REGION Network 9: No encoder pulse
   RUNG wire#powerrail
      Contact( #IN_xFaultsEnabled )
      Contact( #IN_xCycleONDel )
      Contact( #ST_xEncDownPosition )
      { S7_Templates := "SrcType := DInt" } EQ_Contact(in1 := #INPUTS.dEncCounter_count, in2 := #AUX_dLastCounterValueFast_cmm)
      Move(in := #INPUTS.dEncCounter_count, out1 => #AUX_dLastCounterValueFast_cmm)
      Coil( #tALM.tS.xNoEncPulses )
   END_RUNG
   // the same network as SCL:
   #_w1 := #IN_xFaultsEnabled AND #IN_xCycleONDel AND #ST_xEncDownPosition AND (#INPUTS.dEncCounter_count = #AUX_dLastCounterValueFast_cmm);
   IF #_w1 THEN #AUX_dLastCounterValueFast_cmm := #INPUTS.dEncCounter_count; END_IF;
   #tALM.tS.xNoEncPulses := #_w1;
END_REGION

REGION Network 10: Speed values outside limits
   RUNG wire#powerrail
      Contact( #IN_xFaultsEnabled )
      Contact( #IN_xCycleONDel )
      Contact( #ST_xEncDownPosition )
      wire#w1
      { S7_Templates := "SrcType := DInt" } LT_Contact(in1 := #tHMR.dActualEncoderSpeed_mm_min, in2 := "DMINLEHRSPEED_MM_MIN")
      wire#w2
      Coil( #tALM.tS.xSpeedOutLimits )
   END_RUNG
   RUNG wire#w1
      { S7_Templates := "SrcType := DInt" } GT_Contact(in1 := #tHMR.dActualEncoderSpeed_mm_min, in2 := "DMAXLEHRSPEED_MM_MIN")
   END_RUNG wire#w2
   // the same network as SCL:
   #tALM.tS.xSpeedOutLimits := #IN_xFaultsEnabled AND #IN_xCycleONDel AND #ST_xEncDownPosition AND ((#tHMR.dActualEncoderSpeed_mm_min < "DMINLEHRSPEED_MM_MIN") OR (#tHMR.dActualEncoderSpeed_mm_min > "DMAXLEHRSPEED_MM_MIN"));
END_REGION

REGION Network 11: Fm152. Sending data error
   RUNG wire#powerrail
      Contact( #tPhases.xEndPrepareTelegram )
      Contact( #FB_TSend.ERROR )
      S_Coil( #tALM.tF.xFm152SendError )
   END_RUNG
   // the same network as SCL:
   IF #tPhases.xEndPrepareTelegram AND #FB_TSend.ERROR THEN #tALM.tF.xFm152SendError := TRUE; END_IF;
END_REGION

REGION Network 12: FM152.Send data timeout
   #tmON_TimeoutSendData(IN := #tPhases.xPrepareTelegram, PT := #CONST_DTIMEOUTSENDDATA_MS);   // TON
   IF #tmON_TimeoutSendData.Q THEN #tALM.tF.xFm152SendTimeout := TRUE; END_IF;
END_REGION

REGION Network 13: Receive timeout
   #tmON_TimeoutRecvData(IN := #tPhases.xWaitingFm152Reply, PT := #CONST_DTIMEOUTRECVDATA_MS);   // TON
   IF #tmON_TimeoutRecvData.Q THEN
       #tALM.tF.xFm152RecvTimeout := TRUE;
       #AUX_dActualElBuffer := 0;
   END_IF;
END_REGION

REGION Network 14 (SCL): Calculate general statuses
   GATHER(IN:=#tALM.tS,
          OUT=>#TMP_dwValue);

   IF #TMP_dwValue <> 0 THEN
       #ST_xStoppingFaults := TRUE;
   ELSE
       #ST_xStoppingFaults := FALSE;
   END_IF;

   GATHER(IN:=#tALM.tF,
          OUT=>#TMP_dwValue);

   IF #TMP_dwValue <> 0 THEN
       #ST_xFaults := TRUE;
   ELSE
       #ST_xFaults := FALSE;
   END_IF;

   GATHER(IN:=#tALM.tW,
          OUT=>#TMP_dwValue);

   IF #TMP_dwValue <> 0 THEN
       #ST_xWarnings := TRUE;
   ELSE
       #ST_xWarnings := FALSE;
   END_IF;
END_REGION

REGION Network 15: ####_HMI_LOGICS_####
END_REGION

REGION Network 16 (SCL): Manage HMI request
   (*REGION Enable disable glass sensor

       IF #tHMW.xEnableGlassSensor THEN
           #tHMR.xGlassSensorEnabled := TRUE;
           #tHMW.xEnableGlassSensor := FALSE;
       END_IF;

       IF #tHMW.xDisableGlassSensor THEN
           #tHMR.xGlassSensorEnabled := FALSE;
           #tHMW.xDisableGlassSensor := FALSE;
       END_IF;

   END_REGION *)

   REGION Length calibration

       IF #tHMW.xCalibRequest THEN

           #TMP_rF1Unit := DINT_TO_REAL(#tHMW.dCalibRealLength_cmm) / (DINT_TO_REAL(#tHMW.dCalibTheoLength_cmm) / DINT_TO_REAL(#tHMR.dCalibrationF1Unit_unit));
           #tHMR.dCalibrationF1Unit_unit := REAL_TO_DINT(#TMP_rF1Unit);

           #tHMW.dCalibRealLength_cmm := #tHMW.dCalibTheoLength_cmm;        

           #tHMW.xCalibRequest := FALSE;

       END_IF;

   END_REGION

   REGION Update F1

       IF #tHMW.xCalibUpdateF1 THEN

           #tHMR.dCalibrationF1Unit_unit := #tHMW.dCalibWriteF1_unit;
           #tHMW.xCalibUpdateF1 := FALSE;
           #ST_xRefreshFM152 := TRUE;

       END_IF;

   END_REGION

   REGION Update F2

       IF #tHMW.xCalibUpdateF2 THEN

           #tHMR.dCalibrationF2Unit_unit := #tHMW.dCalibWriteF2_unit;
           #tHMW.xCalibUpdateF2 := FALSE;
           #ST_xRefreshFM152 := TRUE;

       END_IF;

   END_REGION
END_REGION

REGION Network 17: Manual command enabled
   RUNG wire#powerrail
      Contact( #tHMW.xEnDisManCom )
      Contact( #ST_xCondOkMan )
      wire#w1
      Coil( #tHMR.xManComEn )
   END_RUNG
   RUNG wire#powerrail
      Contact( #tHMR.xManComEn )
      Contact( #tHMW.xEnDisManCom )
   END_RUNG wire#w1
   // the same network as SCL:
   #tHMR.xManComEn := (#tHMW.xEnDisManCom AND #ST_xCondOkMan) OR (#tHMR.xManComEn AND #tHMW.xEnDisManCom);
END_REGION

REGION Network 18: ####_STATUSES_####
END_REGION

REGION Network 19: Output enable
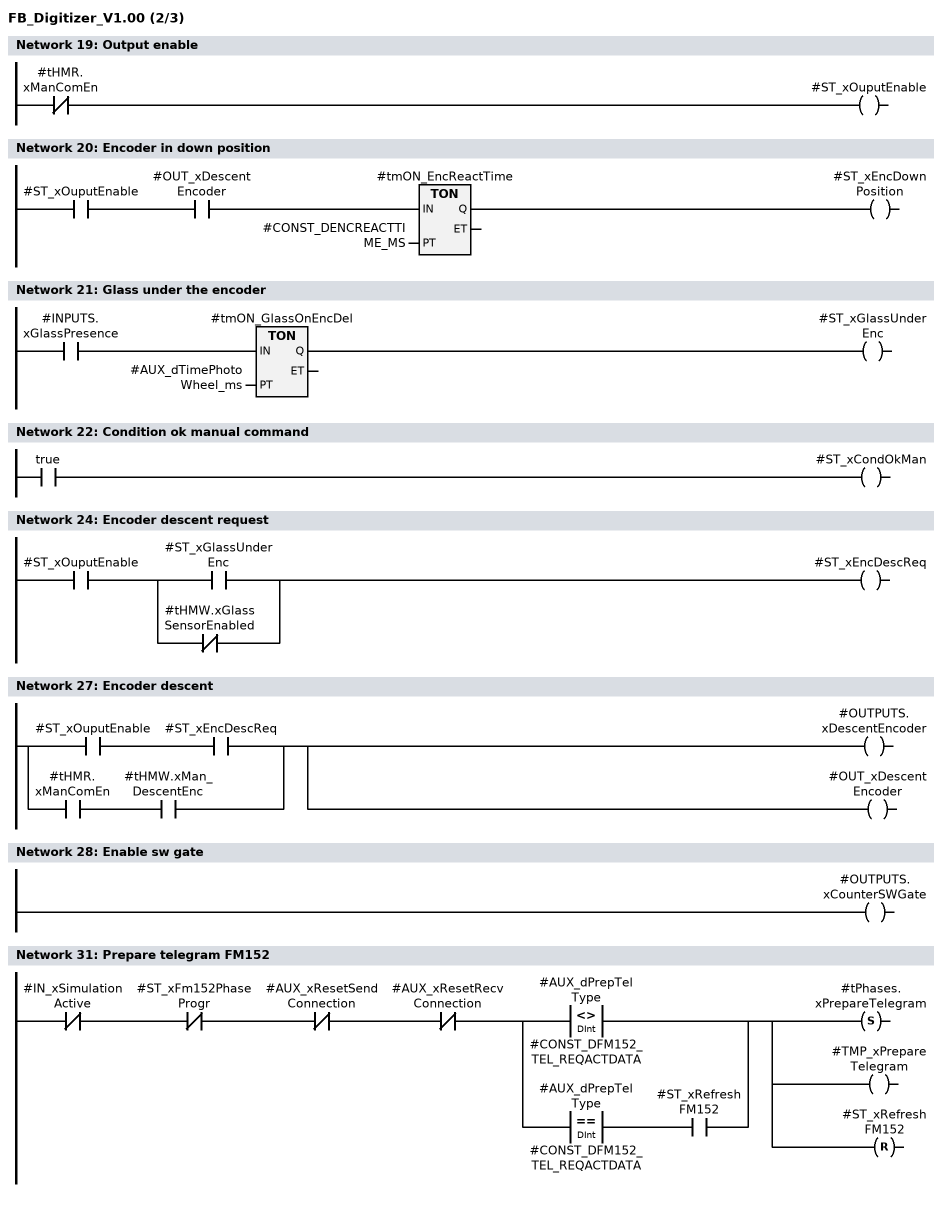
   RUNG wire#powerrail
      I_Contact( #tHMR.xManComEn )
      Coil( #ST_xOuputEnable )
   END_RUNG
   // the same network as SCL:
   #ST_xOuputEnable := NOT #tHMR.xManComEn;
END_REGION

REGION Network 20: Encoder in down position
   #tmON_EncReactTime(IN := #ST_xOuputEnable AND #OUT_xDescentEncoder, PT := #CONST_DENCREACTTIME_MS);   // TON
   #ST_xEncDownPosition := #tmON_EncReactTime.Q;
END_REGION

REGION Network 21: Glass under the encoder
   #tmON_GlassOnEncDel(IN := #INPUTS.xGlassPresence, PT := #AUX_dTimePhotoWheel_ms);   // TON
   #ST_xGlassUnderEnc := #tmON_GlassOnEncDel.Q;
END_REGION

REGION Network 22: Condition ok manual command
   RUNG wire#powerrail
      Contact( true )
      Coil( #ST_xCondOkMan )
   END_RUNG
   // the same network as SCL:
   #ST_xCondOkMan := true;
END_REGION

REGION Network 23: ####_PHASES_&_LOGICS_####
END_REGION

REGION Network 24: Encoder descent request
   RUNG wire#powerrail
      Contact( #ST_xOuputEnable )
      wire#w1
      Contact( #ST_xGlassUnderEnc )
      wire#w2
      Coil( #ST_xEncDescReq )
   END_RUNG
   RUNG wire#w1
      I_Contact( #tHMW.xGlassSensorEnabled )
   END_RUNG wire#w2
   // the same network as SCL:
   #ST_xEncDescReq := #ST_xOuputEnable AND (#ST_xGlassUnderEnc OR NOT #tHMW.xGlassSensorEnabled);
END_REGION

REGION Network 25 (SCL): ####_HMI_STATUSES_####
   #AUX_lrTimingCounter_s += #AUX_lrElapsedTime_s;

   IF #AUX_lrTimingCounter_s >= #CONST_DREFRESHSPEED_S THEN

       #TMP_dElapsedPulses_cmm := #INPUTS.dEncCounter_count - #AUX_dLastCounterValue_cmm;

       #tHMR.dActualEncoderSpeed_mm_min := REAL_TO_DINT(((DINT_TO_REAL(#TMP_dElapsedPulses_cmm) / 100.0) / (LREAL_TO_REAL(#AUX_lrTimingCounter_s))) * 60.0);

       #AUX_dLastCounterValue_cmm := #INPUTS.dEncCounter_count;
       #AUX_lrTimingCounter_s := 0;

   END_IF;

   IF #OUTPUTS.xDescentEncoder AND #tHMW.xMan_DescentEnc THEN
       #tHMR.xMan_DescEncFdbk := TRUE;
   ELSE
       #tHMR.xMan_DescEncFdbk := FALSE;

   END_IF;

   IF #ST_xStoppingFaults THEN
       #tHMR.dEncoderStatus := 7;
   ELSIF #ST_xEncDownPosition THEN
       #tHMR.dEncoderStatus := 3;
   ELSE
       #tHMR.dEncoderStatus := 1;
   END_IF;
END_REGION

REGION Network 26: ####_OUTPUTS_####
END_REGION

REGION Network 27: Encoder descent
   RUNG wire#powerrail
      Contact( #ST_xOuputEnable )
      Contact( #ST_xEncDescReq )
      wire#w1
      Coil( #OUTPUTS.xDescentEncoder )
   END_RUNG
   RUNG wire#powerrail
      Contact( #tHMR.xManComEn )
      Contact( #tHMW.xMan_DescentEnc )
   END_RUNG wire#w1
   RUNG wire#w1
      Coil( #OUT_xDescentEncoder )
   END_RUNG
   // the same network as SCL:
   #OUTPUTS.xDescentEncoder := (#ST_xOuputEnable AND #ST_xEncDescReq) OR (#tHMR.xManComEn AND #tHMW.xMan_DescentEnc);
   #OUT_xDescentEncoder := #OUTPUTS.xDescentEncoder;
END_REGION

REGION Network 28: Enable sw gate
   RUNG wire#powerrail
      Coil( #OUTPUTS.xCounterSWGate )
   END_RUNG
   // the same network as SCL:
   #OUTPUTS.xCounterSWGate := TRUE;
END_REGION

REGION Network 29: ####_ETHERNET_TO_FM152_####
END_REGION

REGION Network 30 (SCL): Initialize connection data
   IF #IN_xGeneralReset THEN

       #AUX_tConnData.InterfaceId := #IN_tInterfaceID;
       #AUX_tConnData.ID := #IN_tID;
       #AUX_tConnData.ConnectionType := #CONST_BCONNTYPE;
       #AUX_tConnData.ActiveEstablished := TRUE;
       #AUX_tConnData.RemoteAddress := #IN_tRemoteAddress;
       #AUX_tConnData.RemotePort := #IN_uiRemotePort;
       #AUX_tConnData.LocalPort := 0;

       //Reset della fasi
       #TMP_dwValue := 0;
       SCATTER(IN:=#TMP_dwValue,
               OUT=>#tPhases);



   END_IF;

   #AUX_xResetRecvConnection := #IN_xGeneralReset;
   #AUX_xResetSendConnection := #IN_xGeneralReset;
END_REGION

REGION Network 31: Prepare telegram FM152
   RUNG wire#powerrail
      I_Contact( #IN_xSimulationActive )
      I_Contact( #ST_xFm152PhaseProgr )
      I_Contact( #AUX_xResetSendConnection )
      I_Contact( #AUX_xResetRecvConnection )
      wire#w1
      { S7_Templates := "SrcType := DInt" } NE_Contact(in1 := #AUX_dPrepTelType, in2 := #CONST_DFM152_TEL_REQACTDATA)
      wire#w2
      S_Coil( #tPhases.xPrepareTelegram )
   END_RUNG
   RUNG wire#w1
      { S7_Templates := "SrcType := DInt" } EQ_Contact(in1 := #AUX_dPrepTelType, in2 := #CONST_DFM152_TEL_REQACTDATA)
      Contact( #ST_xRefreshFM152 )
   END_RUNG wire#w2
   RUNG wire#w2
      Coil( #TMP_xPrepareTelegram )
   END_RUNG
   RUNG wire#w2
      R_Coil( #ST_xRefreshFM152 )
   END_RUNG
   // the same network as SCL:
   #_w1 := NOT #IN_xSimulationActive AND NOT #ST_xFm152PhaseProgr AND NOT #AUX_xResetSendConnection AND NOT #AUX_xResetRecvConnection AND ((#AUX_dPrepTelType <> #CONST_DFM152_TEL_REQACTDATA) OR ((#AUX_dPrepTelType = #CONST_DFM152_TEL_REQACTDATA) AND #ST_xRefreshFM152));
   IF #_w1 THEN #tPhases.xPrepareTelegram := TRUE; END_IF;
   #TMP_xPrepareTelegram := #_w1;
   IF #_w1 THEN #ST_xRefreshFM152 := FALSE; END_IF;
END_REGION

REGION Network 32 (SCL): Prepare telegram
   IF #TMP_xPrepareTelegram THEN

       #AUX_dPrepTelType += 1;

       IF #AUX_dPrepTelType > #CONST_DFM152_TEL_REQACTDATA THEN
           #AUX_dPrepTelType := #CONST_DFM152_TEL_READST;
       END_IF;

       CASE #AUX_dPrepTelType OF

           #CONST_DFM152_TEL_READST:

               #AUX_tFM152SndReadSt.bEOT := #CONST_BFM152_EOT;
               #AUX_tFM152SndReadSt.bAD1 := #CONST_BFM152_AD1;    
               #AUX_tFM152SndReadSt.bAD2 := #CONST_BFM152_AD2;
               #AUX_tFM152SndReadSt.bC1 := '8';
               #AUX_tFM152SndReadSt.bC2 := '5';
               #AUX_tFM152SndReadSt.bENQ := #CONST_BFM152_ENQ;

               #TMP_dBufferPos := 0;
               #TMP_iRetVal := Serialize(SRC_VARIABLE:=#AUX_tFM152SndReadSt, DEST_ARRAY=>#AUX_rgbTempSendBuffer, POS:=#TMP_dBufferPos);
               #AUX_dNumByteToSend := #CONST_DFM152_TEL_READST_NUMBYTE;

           #CONST_DFM152_TEL_READF1:

               #AUX_tFM152SndReadF1.bEOT := #CONST_BFM152_EOT;
               #AUX_tFM152SndReadF1.bAD1 := #CONST_BFM152_AD1;    
               #AUX_tFM152SndReadF1.bAD2 := #CONST_BFM152_AD2;
               #AUX_tFM152SndReadF1.bC1 := '0';
               #AUX_tFM152SndReadF1.bC2 := '0';
               #AUX_tFM152SndReadF1.bENQ := #CONST_BFM152_ENQ;

               #TMP_dBufferPos := 0;
               #TMP_iRetVal := Serialize(SRC_VARIABLE:=#AUX_tFM152SndReadF1, DEST_ARRAY=>#AUX_rgbTempSendBuffer, POS:=#TMP_dBufferPos);
               #AUX_dNumByteToSend := #CONST_DFM152_TEL_READF1_NUMBYTE;

           #CONST_DFM152_TEL_READF2:

               #AUX_tFM152SndReadF2.bEOT := #CONST_BFM152_EOT;
               #AUX_tFM152SndReadF2.bAD1 := #CONST_BFM152_AD1;    
               #AUX_tFM152SndReadF2.bAD2 := #CONST_BFM152_AD2;
               #AUX_tFM152SndReadF2.bC1 := '0';
               #AUX_tFM152SndReadF2.bC2 := '1';
               #AUX_tFM152SndReadF2.bENQ := #CONST_BFM152_ENQ;

               #TMP_dBufferPos := 0;
               #TMP_iRetVal := Serialize(SRC_VARIABLE:=#AUX_tFM152SndReadF2, DEST_ARRAY=>#AUX_rgbTempSendBuffer, POS:=#TMP_dBufferPos);
               #AUX_dNumByteToSend := #CONST_DFM152_TEL_READF2_NUMBYTE;

           #CONST_DFM152_TEL_WRITEF1:

               #TMP_strValue := DINT_TO_STRING(#tHMR.dCalibrationF1Unit_unit);

               #AUX_tFM152SndWriteF1.bEOT := #CONST_BFM152_EOT;
               #AUX_tFM152SndWriteF1.bAD1 := #CONST_BFM152_AD1;
               #AUX_tFM152SndWriteF1.bAD2 := #CONST_BFM152_AD2;
               #AUX_tFM152SndWriteF1.bSTX := #CONST_BFM152_STX;
               #AUX_tFM152SndWriteF1.bC1 := '0';
               #AUX_tFM152SndWriteF1.bC2 := '0';
               #AUX_tFM152SndWriteF1.bVal1 := #TMP_strValue[2];
               #AUX_tFM152SndWriteF1.bVal2 := #TMP_strValue[3];
               #AUX_tFM152SndWriteF1.bVal3 := #TMP_strValue[4];
               #AUX_tFM152SndWriteF1.bVal4 := #TMP_strValue[5];
               #AUX_tFM152SndWriteF1.bVal5 := #TMP_strValue[6];
               #AUX_tFM152SndWriteF1.bETX := #CONST_BFM152_ETX;
               #AUX_tFM152SndWriteF1.bBCC := #AUX_tFM152SndWriteF1.bC1; 
               #AUX_tFM152SndWriteF1.bBCC := #AUX_tFM152SndWriteF1.bBCC XOR #AUX_tFM152SndWriteF1.bC2;
               #AUX_tFM152SndWriteF1.bBCC := #AUX_tFM152SndWriteF1.bBCC XOR #AUX_tFM152SndWriteF1.bVal1;
               #AUX_tFM152SndWriteF1.bBCC := #AUX_tFM152SndWriteF1.bBCC XOR #AUX_tFM152SndWriteF1.bVal2;
               #AUX_tFM152SndWriteF1.bBCC := #AUX_tFM152SndWriteF1.bBCC XOR #AUX_tFM152SndWriteF1.bVal3;
               #AUX_tFM152SndWriteF1.bBCC := #AUX_tFM152SndWriteF1.bBCC XOR #AUX_tFM152SndWriteF1.bVal4;
               #AUX_tFM152SndWriteF1.bBCC := #AUX_tFM152SndWriteF1.bBCC XOR #AUX_tFM152SndWriteF1.bVal5;
               #AUX_tFM152SndWriteF1.bBCC := #AUX_tFM152SndWriteF1.bBCC XOR #AUX_tFM152SndWriteF1.bETX; 

               #TMP_dBufferPos := 0;
               #TMP_iRetVal := Serialize(SRC_VARIABLE:=#AUX_tFM152SndWriteF1, DEST_ARRAY=>#AUX_rgbTempSendBuffer, POS:=#TMP_dBufferPos);
               #AUX_dNumByteToSend := #CONST_DFM152_TEL_WRITEF1_NUMBYTE;

           #CONST_DFM152_TEL_WRITEF2:

               #TMP_strValue := DINT_TO_STRING(#tHMR.dCalibrationF2Unit_unit);

               #AUX_tFM152SndWriteF2.bEOT := #CONST_BFM152_EOT;
               #AUX_tFM152SndWriteF2.bAD1 := #CONST_BFM152_AD1;
               #AUX_tFM152SndWriteF2.bAD2 := #CONST_BFM152_AD2;
               #AUX_tFM152SndWriteF2.bSTX := #CONST_BFM152_STX;
               #AUX_tFM152SndWriteF2.bC1 := '0';
               #AUX_tFM152SndWriteF2.bC2 := '1';
               #AUX_tFM152SndWriteF2.bVal1 := #TMP_strValue[2];
               #AUX_tFM152SndWriteF2.bVal2 := #TMP_strValue[3];
               #AUX_tFM152SndWriteF2.bVal3 := #TMP_strValue[4];
               #AUX_tFM152SndWriteF2.bVal4 := #TMP_strValue[5];
               #AUX_tFM152SndWriteF2.bVal5 := #TMP_strValue[6];
               #AUX_tFM152SndWriteF2.bETX := #CONST_BFM152_ETX;
               #AUX_tFM152SndWriteF2.bBCC := #AUX_tFM152SndWriteF2.bC1; 
               #AUX_tFM152SndWriteF2.bBCC := #AUX_tFM152SndWriteF2.bBCC XOR #AUX_tFM152SndWriteF2.bC2;
               #AUX_tFM152SndWriteF2.bBCC := #AUX_tFM152SndWriteF2.bBCC XOR #AUX_tFM152SndWriteF2.bVal1;
               #AUX_tFM152SndWriteF2.bBCC := #AUX_tFM152SndWriteF2.bBCC XOR #AUX_tFM152SndWriteF2.bVal2;
               #AUX_tFM152SndWriteF2.bBCC := #AUX_tFM152SndWriteF2.bBCC XOR #AUX_tFM152SndWriteF2.bVal3;
               #AUX_tFM152SndWriteF2.bBCC := #AUX_tFM152SndWriteF2.bBCC XOR #AUX_tFM152SndWriteF2.bVal4;
               #AUX_tFM152SndWriteF2.bBCC := #AUX_tFM152SndWriteF2.bBCC XOR #AUX_tFM152SndWriteF2.bVal5;
               #AUX_tFM152SndWriteF2.bBCC := #AUX_tFM152SndWriteF2.bBCC XOR #AUX_tFM152SndWriteF2.bETX; 

               #TMP_dBufferPos := 0;
               #TMP_iRetVal := Serialize(SRC_VARIABLE:=#AUX_tFM152SndWriteF2, DEST_ARRAY=>#AUX_rgbTempSendBuffer, POS:=#TMP_dBufferPos);
               #AUX_dNumByteToSend := #CONST_DFM152_TEL_WRITEF2_NUMBYTE;

           #CONST_DFM152_TEL_WRITEJOG:

               #TMP_strValue := DINT_TO_STRING(REAL_TO_DINT((DINT_TO_REAL(#tHMW.dRequestJogSpeed_mm_min) * 100.0) / 60.0));
               #AUX_tFM152SndWriteJog.bEOT := #CONST_BFM152_EOT;
               #AUX_tFM152SndWriteJog.bAD1 := #CONST_BFM152_AD1;
               #AUX_tFM152SndWriteJog.bAD2 :=  #CONST_BFM152_AD2;
               #AUX_tFM152SndWriteJog.bSTX := #CONST_BFM152_STX;
               #AUX_tFM152SndWriteJog.bC1 := '0'; 
               #AUX_tFM152SndWriteJog.bC2 := '5'; 
               #AUX_tFM152SndWriteJog.bVal1 := #TMP_strValue[2];
               #AUX_tFM152SndWriteJog.bVal2 := #TMP_strValue[3];
               #AUX_tFM152SndWriteJog.bVal3 := #TMP_strValue[4];
               #AUX_tFM152SndWriteJog.bVal4 := #TMP_strValue[5];
               #AUX_tFM152SndWriteJog.bVal5 := #TMP_strValue[6];
               #AUX_tFM152SndWriteJog.bETX := #CONST_BFM152_ETX;
               #AUX_tFM152SndWriteJog.bBCC := #AUX_tFM152SndWriteJog.bC1; 
               #AUX_tFM152SndWriteJog.bBCC := #AUX_tFM152SndWriteJog.bBCC XOR #AUX_tFM152SndWriteJog.bC2;
               #AUX_tFM152SndWriteJog.bBCC := #AUX_tFM152SndWriteJog.bBCC XOR #AUX_tFM152SndWriteJog.bVal1;
               #AUX_tFM152SndWriteJog.bBCC := #AUX_tFM152SndWriteJog.bBCC XOR #AUX_tFM152SndWriteJog.bVal2;
               #AUX_tFM152SndWriteJog.bBCC := #AUX_tFM152SndWriteJog.bBCC XOR #AUX_tFM152SndWriteJog.bVal3;
               #AUX_tFM152SndWriteJog.bBCC := #AUX_tFM152SndWriteJog.bBCC XOR #AUX_tFM152SndWriteJog.bVal4;
               #AUX_tFM152SndWriteJog.bBCC := #AUX_tFM152SndWriteJog.bBCC XOR #AUX_tFM152SndWriteJog.bVal5;
               #AUX_tFM152SndWriteJog.bBCC := #AUX_tFM152SndWriteJog.bBCC XOR #AUX_tFM152SndWriteJog.bETX;

               #TMP_dBufferPos := 0;
               #TMP_iRetVal := Serialize(SRC_VARIABLE:=#AUX_tFM152SndWriteJog, DEST_ARRAY=>#AUX_rgbTempSendBuffer, POS:=#TMP_dBufferPos);
               #AUX_dNumByteToSend := #CONST_DFM152_TEL_WRITEJOG_NUMBYTE;


           #CONST_DFM152_TEL_WRITERAMPREF:

               #AUX_tFM152SndWriteRampRef.bEOT := #CONST_BFM152_EOT;
               #AUX_tFM152SndWriteRampRef.bAD1 := #CONST_BFM152_AD1;
               #AUX_tFM152SndWriteRampRef.bAD2 := #CONST_BFM152_AD2;
               #AUX_tFM152SndWriteRampRef.bSTX := #CONST_BFM152_STX;
               #AUX_tFM152SndWriteRampRef.bC1 := '0';
               #AUX_tFM152SndWriteRampRef.bC2 := '4';
               #AUX_tFM152SndWriteRampRef.bC3 := '0';
               #AUX_tFM152SndWriteRampRef.bC4 := '0';
               #AUX_tFM152SndWriteRampRef.bETX := #CONST_BFM152_ETX;
               #AUX_tFM152SndWriteRampRef.bBCC := #AUX_tFM152SndWriteRampRef.bC1;
               #AUX_tFM152SndWriteRampRef.bBCC :=  #AUX_tFM152SndWriteRampRef.bBCC XOR #AUX_tFM152SndWriteRampRef.bC2;
               #AUX_tFM152SndWriteRampRef.bBCC :=  #AUX_tFM152SndWriteRampRef.bBCC XOR #AUX_tFM152SndWriteRampRef.bC3;
               #AUX_tFM152SndWriteRampRef.bBCC :=  #AUX_tFM152SndWriteRampRef.bBCC XOR #AUX_tFM152SndWriteRampRef.bC4;
               #AUX_tFM152SndWriteRampRef.bBCC :=  #AUX_tFM152SndWriteRampRef.bBCC XOR #AUX_tFM152SndWriteRampRef.bETX;

               #TMP_dBufferPos := 0;
               #TMP_iRetVal := Serialize(SRC_VARIABLE:=#AUX_tFM152SndWriteRampRef, DEST_ARRAY=>#AUX_rgbTempSendBuffer, POS:=#TMP_dBufferPos);
               #AUX_dNumByteToSend := #CONST_DFM152_TEL_WRITERAMPREF_NUMBYTE;


           #CONST_DFM152_TEL_WRITERAMPJOG:

               #AUX_tFM152SndWriteRampJog.bEOT := #CONST_BFM152_EOT;
               #AUX_tFM152SndWriteRampJog.bAD1 := #CONST_BFM152_AD1;
               #AUX_tFM152SndWriteRampJog.bAD2 := #CONST_BFM152_AD2;
               #AUX_tFM152SndWriteRampJog.bSTX := #CONST_BFM152_STX;
               #AUX_tFM152SndWriteRampJog.bC1 := '0';
               #AUX_tFM152SndWriteRampJog.bC2 := '6';
               #AUX_tFM152SndWriteRampJog.bC3 := '0';
               #AUX_tFM152SndWriteRampJog.bC4 := '0';
               #AUX_tFM152SndWriteRampJog.bETX := #CONST_BFM152_ETX;
               #AUX_tFM152SndWriteRampJog.bBCC := #AUX_tFM152SndWriteRampJog.bC1;
               #AUX_tFM152SndWriteRampJog.bBCC := #AUX_tFM152SndWriteRampJog.bBCC XOR #AUX_tFM152SndWriteRampJog.bC2;
               #AUX_tFM152SndWriteRampJog.bBCC := #AUX_tFM152SndWriteRampJog.bBCC XOR #AUX_tFM152SndWriteRampJog.bC3;
               #AUX_tFM152SndWriteRampJog.bBCC := #AUX_tFM152SndWriteRampJog.bBCC XOR #AUX_tFM152SndWriteRampJog.bC4;
               #AUX_tFM152SndWriteRampJog.bBCC := #AUX_tFM152SndWriteRampJog.bBCC XOR #AUX_tFM152SndWriteRampJog.bETX;

               #TMP_dBufferPos := 0;
               #TMP_iRetVal := Serialize(SRC_VARIABLE:=#AUX_tFM152SndWriteRampJog, DEST_ARRAY=>#AUX_rgbTempSendBuffer, POS:=#TMP_dBufferPos);
               #AUX_dNumByteToSend := #CONST_DFM152_TEL_WRITERAMPJOG_NUMBYTE;

           #CONST_DFM152_TEL_WRITERAMP:

               #AUX_tFM152SndWriteRamp.bEOT := #CONST_BFM152_EOT;
               #AUX_tFM152SndWriteRamp.bAD1 := #CONST_BFM152_AD1;
               #AUX_tFM152SndWriteRamp.bAD2 := #CONST_BFM152_AD2;
               #AUX_tFM152SndWriteRamp.bSTX := #CONST_BFM152_STX;
               #AUX_tFM152SndWriteRamp.bC1 := '0';
               #AUX_tFM152SndWriteRamp.bC2 := '9';
               #AUX_tFM152SndWriteRamp.bC3 := '0';
               #AUX_tFM152SndWriteRamp.bC4 := '0';
               #AUX_tFM152SndWriteRamp.bETX := #CONST_BFM152_ETX;
               #AUX_tFM152SndWriteRamp.bBCC := #AUX_tFM152SndWriteRamp.bC1;
               #AUX_tFM152SndWriteRamp.bBCC := #AUX_tFM152SndWriteRamp.bBCC XOR #AUX_tFM152SndWriteRamp.bC2;
               #AUX_tFM152SndWriteRamp.bBCC := #AUX_tFM152SndWriteRamp.bBCC XOR #AUX_tFM152SndWriteRamp.bC3;
               #AUX_tFM152SndWriteRamp.bBCC := #AUX_tFM152SndWriteRamp.bBCC XOR #AUX_tFM152SndWriteRamp.bC4;
               #AUX_tFM152SndWriteRamp.bBCC := #AUX_tFM152SndWriteRamp.bBCC XOR #AUX_tFM152SndWriteRamp.bETX;

               #TMP_dBufferPos := 0;
               #TMP_iRetVal := Serialize(SRC_VARIABLE:=#AUX_tFM152SndWriteRamp, DEST_ARRAY=>#AUX_rgbTempSendBuffer, POS:=#TMP_dBufferPos);
               #AUX_dNumByteToSend := #CONST_DFM152_TEL_WRITERAMP_NUMBYTE;


           #CONST_DFM152_TEL_REQACTDATA:

               #AUX_tFM152SndActivateData.bEOT := #CONST_BFM152_EOT;
               #AUX_tFM152SndActivateData.bAD1 := #CONST_BFM152_AD1;
               #AUX_tFM152SndActivateData.bAD2 := #CONST_BFM152_AD2;
               #AUX_tFM152SndActivateData.bSTX := #CONST_BFM152_STX;
               #AUX_tFM152SndActivateData.bC1 := '6';
               #AUX_tFM152SndActivateData.bC2 := '7';
               #AUX_tFM152SndActivateData.bC3 := '1';
               #AUX_tFM152SndActivateData.bETX := #CONST_BFM152_ETX;
               #AUX_tFM152SndActivateData.bBCC := #AUX_tFM152SndActivateData.bC1;
               #AUX_tFM152SndActivateData.bBCC := #AUX_tFM152SndActivateData.bBCC XOR #AUX_tFM152SndActivateData.bC2;
               #AUX_tFM152SndActivateData.bBCC := #AUX_tFM152SndActivateData.bBCC XOR #AUX_tFM152SndActivateData.bC3;
               #AUX_tFM152SndActivateData.bBCC := #AUX_tFM152SndActivateData.bBCC XOR #AUX_tFM152SndActivateData.bETX;

               #TMP_dBufferPos := 0;
               #TMP_iRetVal := Serialize(SRC_VARIABLE:=#AUX_tFM152SndActivateData, DEST_ARRAY=>#AUX_rgbTempSendBuffer, POS:=#TMP_dBufferPos);
               #AUX_dNumByteToSend := #CONST_DFM152_TEL_REQACTDATA_NUMBYTE;

       END_CASE;
   END_IF;
END_REGION

REGION Network 33: ### SEND DATA TO FM
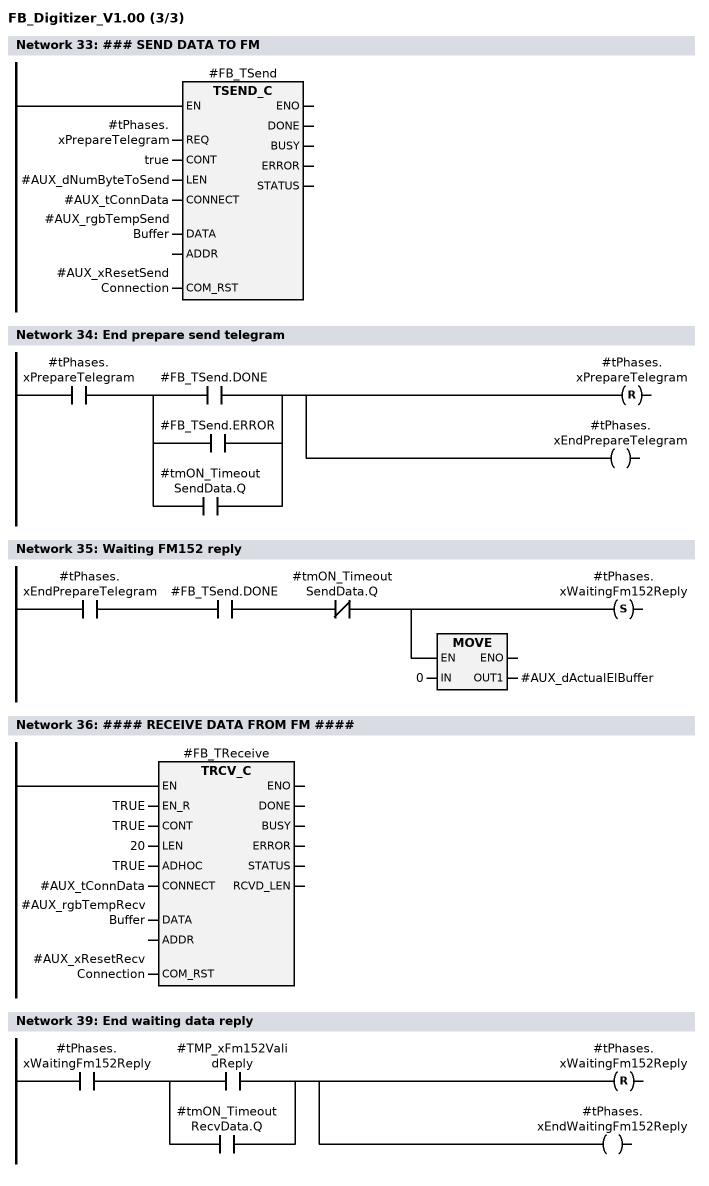
   #FB_TSend(REQ := #tPhases.xPrepareTelegram,   // TSEND_C
             CONT := true,
             LEN := #AUX_dNumByteToSend,
             CONNECT := #AUX_tConnData,
             DATA := #AUX_rgbTempSendBuffer,
             COM_RST := #AUX_xResetSendConnection);
END_REGION

REGION Network 34: End prepare send telegram
   RUNG wire#powerrail
      Contact( #tPhases.xPrepareTelegram )
      wire#w1
      Contact( #FB_TSend.DONE )
      wire#w2
      R_Coil( #tPhases.xPrepareTelegram )
   END_RUNG
   RUNG wire#w1
      Contact( #FB_TSend.ERROR )
   END_RUNG wire#w2
   RUNG wire#w1
      Contact( #tmON_TimeoutSendData.Q )
   END_RUNG wire#w2
   RUNG wire#w2
      Coil( #tPhases.xEndPrepareTelegram )
   END_RUNG
   // the same network as SCL:
   #_w1 := #tPhases.xPrepareTelegram AND (#FB_TSend.DONE OR #FB_TSend.ERROR OR #tmON_TimeoutSendData.Q);
   IF #_w1 THEN #tPhases.xPrepareTelegram := FALSE; END_IF;
   #tPhases.xEndPrepareTelegram := #_w1;
END_REGION

REGION Network 35: Waiting FM152 reply
   RUNG wire#powerrail
      Contact( #tPhases.xEndPrepareTelegram )
      Contact( #FB_TSend.DONE )
      I_Contact( #tmON_TimeoutSendData.Q )
      wire#w1
      S_Coil( #tPhases.xWaitingFm152Reply )
   END_RUNG
   RUNG wire#w1
      Move(in := 0, out1 => #AUX_dActualElBuffer)
   END_RUNG
   // the same network as SCL:
   IF #tPhases.xEndPrepareTelegram AND #FB_TSend.DONE AND NOT #tmON_TimeoutSendData.Q THEN
       #tPhases.xWaitingFm152Reply := TRUE;
       #AUX_dActualElBuffer := 0;
   END_IF;
END_REGION

REGION Network 36: #### RECEIVE DATA FROM FM ####
   #FB_TReceive(EN_R := TRUE,   // TRCV_C
                CONT := TRUE,
                LEN := 20,
                ADHOC := TRUE,
                CONNECT := #AUX_tConnData,
                DATA := #AUX_rgbTempRecvBuffer,
                COM_RST := #AUX_xResetRecvConnection);
END_REGION

REGION Network 37 (SCL): Manage data received
   IF #FB_TReceive.DONE THEN

       IF #FB_TReceive.RCVD_LEN > 0 THEN

           //Copy the byte received from the temp buffer to the destination buffer
           IF (#AUX_dActualElBuffer + UDINT_TO_DINT(#FB_TReceive.RCVD_LEN)) >= 20 THEN
               #AUX_dActualElBuffer := 0;
           END_IF;

           MOVE_BLK(IN:=#AUX_rgbTempRecvBuffer[0],
                    COUNT:=#FB_TReceive.LEN,
                    OUT=>#AUX_rgbReceiveBuffer[#AUX_dActualElBuffer]);

           #AUX_dActualElBuffer+= UDINT_TO_DINT(#FB_TReceive.RCVD_LEN);

       END_IF;

   END_IF;
END_REGION

REGION Network 38 (SCL): Checking the received buffer
   #TMP_xFm152ValidReply := FALSE;

   IF #tPhases.xWaitingFm152Reply THEN

       CASE #AUX_dPrepTelType OF

           #CONST_DFM152_TEL_READST: 

               IF #AUX_dActualElBuffer = #CONST_DFM152_RECVSTATUSSIZE THEN

                   #TMP_dBufferPos := 0;
                   #TMP_iRetVal := Deserialize(SRC_ARRAY:=#AUX_rgbReceiveBuffer, DEST_VARIABLE=>#AUX_tFM152RecvStatus, POS:=#TMP_dBufferPos);

                   //Calculate BCC
                   #TMP_bBBC := #AUX_tFM152RecvStatus.bC1;
                   #TMP_bBBC := #TMP_bBBC XOR #AUX_tFM152RecvStatus.bC2;
                   #TMP_bBBC := #TMP_bBBC XOR #AUX_tFM152RecvStatus.bC3;
                   #TMP_bBBC := #TMP_bBBC XOR #AUX_tFM152RecvStatus.bC4;
                   #TMP_bBBC := #TMP_bBBC XOR #AUX_tFM152RecvStatus.bC5;
                   #TMP_bBBC := #TMP_bBBC XOR #AUX_tFM152RecvStatus.bD1;
                   #TMP_bBBC := #TMP_bBBC XOR #AUX_tFM152RecvStatus.bD2;
                   #TMP_bBBC := #TMP_bBBC XOR #AUX_tFM152RecvStatus.bETX;

                   IF  #AUX_tFM152RecvStatus.bSTX = #CONST_BFM152_STX AND
                       #AUX_tFM152RecvStatus.bC1 = '8' AND
                       #AUX_tFM152RecvStatus.bC2 = '5' AND
                       #AUX_tFM152RecvStatus.bC3 = 'H' AND
                       #AUX_tFM152RecvStatus.bC4 = '0' AND
                       #AUX_tFM152RecvStatus.bC5 = '0' AND
                       #AUX_tFM152RecvStatus.bETX = #CONST_BFM152_ETX AND
                       #AUX_tFM152RecvStatus.bBCC = #TMP_bBBC THEN

                           //Copy the status values
                           #TMP_strStatus[1] := #AUX_tFM152RecvStatus.bD1;
                           #TMP_strStatus[2] := #AUX_tFM152RecvStatus.bD2;

                           #tHMR.dFm152Status := STRING_TO_DINT(#TMP_strStatus);                                  

                           #TMP_xFm152ValidReply := TRUE;
                   END_IF;



               END_IF;

           #CONST_DFM152_TEL_READF1: 

               IF #AUX_dActualElBuffer = #CONST_DFM152_RECVF1F2SIZE THEN

                   #TMP_dBufferPos := 0;
                   #TMP_iRetVal := Deserialize(SRC_ARRAY:=#AUX_rgbReceiveBuffer, DEST_VARIABLE=>#AUX_tFM152RecvF1, POS:=#TMP_dBufferPos);

                   //Calculate BCC
                   #TMP_bBBC :=    #AUX_tFM152RecvF1.bC1;
                   #TMP_bBBC :=    #TMP_bBBC XOR #AUX_tFM152RecvF1.bC2; 
                   #TMP_bBBC :=    #TMP_bBBC XOR #AUX_tFM152RecvF1.bD1; 
                   #TMP_bBBC :=    #TMP_bBBC XOR #AUX_tFM152RecvF1.bD2; 
                   #TMP_bBBC :=    #TMP_bBBC XOR #AUX_tFM152RecvF1.bD3;
                   #TMP_bBBC :=    #TMP_bBBC XOR #AUX_tFM152RecvF1.bD4; 
                   #TMP_bBBC :=    #TMP_bBBC XOR #AUX_tFM152RecvF1.bD5; 
                   #TMP_bBBC :=    #TMP_bBBC XOR #AUX_tFM152RecvF1.bETX;

                   IF  #AUX_tFM152RecvF1.bSTX = #CONST_BFM152_STX AND
                       #AUX_tFM152RecvF1.bC1 = '0' AND
                       #AUX_tFM152RecvF1.bC2 = '0' AND
                       #AUX_tFM152RecvF1.bETX = #CONST_BFM152_ETX AND
                       #AUX_tFM152RecvF1.bBCC = #TMP_bBBC THEN

                           #TMP_strF1F2Value[1] := #AUX_tFM152RecvF1.bD1;
                           #TMP_strF1F2Value[2] := #AUX_tFM152RecvF1.bD2;
                           #TMP_strF1F2Value[3] := #AUX_tFM152RecvF1.bD3;
                           #TMP_strF1F2Value[4] := #AUX_tFM152RecvF1.bD4;
                           #TMP_strF1F2Value[5] := #AUX_tFM152RecvF1.bD5;

                           #tHMR.dCalibrationCardF1Unit_unit := STRING_TO_DINT(#TMP_strF1F2Value);

                           #TMP_xFm152ValidReply := TRUE;    
                   END_IF;

               END_IF;

           #CONST_DFM152_TEL_READF2: 

               IF #AUX_dActualElBuffer = #CONST_DFM152_RECVF1F2SIZE THEN

                   #TMP_dBufferPos := 0;
                   #TMP_iRetVal := Deserialize(SRC_ARRAY:=#AUX_rgbReceiveBuffer, DEST_VARIABLE=>#AUX_tFM152RecvF2, POS:=#TMP_dBufferPos);

                   //Calculate BCC
                   #TMP_bBBC := #AUX_tFM152RecvF2.bC1;
                   #TMP_bBBC := #TMP_bBBC XOR #AUX_tFM152RecvF2.bC2; 
                   #TMP_bBBC := #TMP_bBBC XOR #AUX_tFM152RecvF2.bD1; 
                   #TMP_bBBC := #TMP_bBBC XOR #AUX_tFM152RecvF2.bD2; 
                   #TMP_bBBC := #TMP_bBBC XOR #AUX_tFM152RecvF2.bD3;
                   #TMP_bBBC := #TMP_bBBC XOR #AUX_tFM152RecvF2.bD4; 
                   #TMP_bBBC := #TMP_bBBC XOR #AUX_tFM152RecvF2.bD5; 
                   #TMP_bBBC := #TMP_bBBC XOR #AUX_tFM152RecvF2.bETX;

                   IF  #AUX_tFM152RecvF2.bSTX = #CONST_BFM152_STX AND
                       #AUX_tFM152RecvF2.bC1 = '0' AND
                       #AUX_tFM152RecvF2.bC2 = '1' AND
                       #AUX_tFM152RecvF2.bETX = #CONST_BFM152_ETX AND
                       #AUX_tFM152RecvF2.bBCC = #TMP_bBBC THEN

                           #TMP_strF1F2Value[1] := #AUX_tFM152RecvF2.bD1;
                           #TMP_strF1F2Value[2] := #AUX_tFM152RecvF2.bD2;
                           #TMP_strF1F2Value[3] := #AUX_tFM152RecvF2.bD3;
                           #TMP_strF1F2Value[4] := #AUX_tFM152RecvF2.bD4;
                           #TMP_strF1F2Value[5] := #AUX_tFM152RecvF2.bD5;

                           #tHMR.dCalibrationCardF2Unit_unit := STRING_TO_DINT(#TMP_strF1F2Value);

                           #TMP_xFm152ValidReply := TRUE;    
                   END_IF;

               END_IF;

           #CONST_DFM152_TEL_WRITEF1:        

               IF #AUX_dActualElBuffer = #CONST_DFM152_ACK_NACKSIZE THEN

                   #TMP_dBufferPos := 0;
                   #TMP_iRetVal := Deserialize(SRC_ARRAY:=#AUX_rgbReceiveBuffer, DEST_VARIABLE=>#AUX_tFM152RecvAck, POS:=#TMP_dBufferPos);

                   IF #AUX_tFM152RecvAck.bACK = #CONST_BFM152_ACK THEN
                       #TMP_xFm152ValidReply := TRUE;
                   END_IF;
               END_IF;

           #CONST_DFM152_TEL_WRITEF2:        

               IF #AUX_dActualElBuffer = #CONST_DFM152_ACK_NACKSIZE THEN

                   #TMP_dBufferPos := 0;
                   #TMP_iRetVal := Deserialize(SRC_ARRAY:=#AUX_rgbReceiveBuffer, DEST_VARIABLE=>#AUX_tFM152RecvAck, POS:=#TMP_dBufferPos);

                   IF #AUX_tFM152RecvAck.bACK = #CONST_BFM152_ACK THEN
                       #TMP_xFm152ValidReply := TRUE;
                   END_IF;
               END_IF;

           #CONST_DFM152_TEL_WRITEJOG:        

               IF #AUX_dActualElBuffer = #CONST_DFM152_ACK_NACKSIZE THEN

                   #TMP_dBufferPos := 0;
                   #TMP_iRetVal := Deserialize(SRC_ARRAY:=#AUX_rgbReceiveBuffer, DEST_VARIABLE=>#AUX_tFM152RecvAck, POS:=#TMP_dBufferPos);

                   IF #AUX_tFM152RecvAck.bACK = #CONST_BFM152_ACK THEN
                       #TMP_xFm152ValidReply := TRUE;
                   END_IF;
               END_IF;

           #CONST_DFM152_TEL_WRITERAMPREF:        

               IF #AUX_dActualElBuffer = #CONST_DFM152_ACK_NACKSIZE THEN

                   #TMP_dBufferPos := 0;
                   #TMP_iRetVal := Deserialize(SRC_ARRAY:=#AUX_rgbReceiveBuffer, DEST_VARIABLE=>#AUX_tFM152RecvAck, POS:=#TMP_dBufferPos);